HMI tags "xDI"
   "DIx_DB_M1_QF_Input" : Bool = PLC DIx_DB.M1_QF.Input AT %DB200.DBX0.0, 1 s
   "DIx_DB_M1_QF_Signal" : Bool = PLC DIx_DB.M1_QF.Signal AT %DB200.DBX2.0, 1 s
   "DIx_DB_M1_QF_Hand" : Bool = PLC DIx_DB.M1_QF.Hand AT %DB200.DBX4.0, 1 s
   "DIx_DB_M1_QF_Start_M" : Bool = PLC DIx_DB.M1_QF.Start_M AT %DB200.DBX4.1, 1 s
   "DIx_DB_M1_QF_Inverse" : Bool = PLC DIx_DB.M1_QF.Inverse AT %DB200.DBX4.3, 1 s
   "DIx_DB_M1_QF_Filter_On_SP" : Int = PLC DIx_DB.M1_QF.Filter_On.SP AT %DB200.DBW6, 1 s
   "DIx_DB_M1_QF_Filter_Off_SP" : Int = PLC DIx_DB.M1_QF.Filter_Off.SP AT %DB200.DBW12, 1 s
   "DIx_DB_M2_QF_Input" : Bool = PLC DIx_DB.M2_QF.Input AT %DB200.DBX20.0, 1 s
   "DIx_DB_M2_QF_Signal" : Bool = PLC DIx_DB.M2_QF.Signal AT %DB200.DBX22.0, 1 s
   "DIx_DB_M2_QF_Hand" : Bool = PLC DIx_DB.M2_QF.Hand AT %DB200.DBX24.0, 1 s
   "DIx_DB_M2_QF_Start_M" : Bool = PLC DIx_DB.M2_QF.Start_M AT %DB200.DBX24.1, 1 s
   "DIx_DB_M2_QF_Inverse" : Bool = PLC DIx_DB.M2_QF.Inverse AT %DB200.DBX24.3, 1 s
   "DIx_DB_M2_QF_Filter_On_SP" : Int = PLC DIx_DB.M2_QF.Filter_On.SP AT %DB200.DBW26, 1 s
   "DIx_DB_M2_QF_Filter_Off_SP" : Int = PLC DIx_DB.M2_QF.Filter_Off.SP AT %DB200.DBW32, 1 s
   "DIx_DB_M3_QF_Input" : Bool = PLC DIx_DB.M3_QF.Input AT %DB200.DBX40.0, 1 s
   "DIx_DB_M3_QF_Signal" : Bool = PLC DIx_DB.M3_QF.Signal AT %DB200.DBX42.0, 1 s
   "DIx_DB_M3_QF_Hand" : Bool = PLC DIx_DB.M3_QF.Hand AT %DB200.DBX44.0, 1 s
   "DIx_DB_M3_QF_Start_M" : Bool = PLC DIx_DB.M3_QF.Start_M AT %DB200.DBX44.1, 1 s
   "DIx_DB_M3_QF_Inverse" : Bool = PLC DIx_DB.M3_QF.Inverse AT %DB200.DBX44.3, 1 s
   "DIx_DB_M3_QF_Filter_On_SP" : Int = PLC DIx_DB.M3_QF.Filter_On.SP AT %DB200.DBW46, 1 s
   "DIx_DB_M3_QF_Filter_Off_SP" : Int = PLC DIx_DB.M3_QF.Filter_Off.SP AT %DB200.DBW52, 1 s
   "DIx_DB_Heat_1_Input" : Bool = PLC DIx_DB.Heat_1.Input AT %DB200.DBX60.0, 1 s
   "DIx_DB_Heat_1_Signal" : Bool = PLC DIx_DB.Heat_1.Signal AT %DB200.DBX62.0, 1 s
   "DIx_DB_Heat_1_Hand" : Bool = PLC DIx_DB.Heat_1.Hand AT %DB200.DBX64.0, 1 s
   "DIx_DB_Heat_1_Start_M" : Bool = PLC DIx_DB.Heat_1.Start_M AT %DB200.DBX64.1, 1 s
   "DIx_DB_Heat_1_Filter_On_SP" : Int = PLC DIx_DB.Heat_1.Filter_On.SP AT %DB200.DBW66, 1 s
   "DIx_DB_Heat_1_Filter_Off_SP" : Int = PLC DIx_DB.Heat_1.Filter_Off.SP AT %DB200.DBW72, 1 s
   "DIx_DB_Heat_2_Filter_Off_SP" : Int = PLC DIx_DB.Heat_2.Filter_Off.SP AT %DB200.DBW92, 1 s
   "DIx_DB_Heat_2_Filter_On_SP" : Int = PLC DIx_DB.Heat_2.Filter_On.SP AT %DB200.DBW86, 1 s
   "DIx_DB_Heat_2_Inverse" : Bool = PLC DIx_DB.Heat_2.Inverse AT %DB200.DBX84.3, 1 s
   "DIx_DB_Heat_2_Start_M" : Bool = PLC DIx_DB.Heat_2.Start_M AT %DB200.DBX84.1, 1 s
   "DIx_DB_Heat_2_Hand" : Bool = PLC DIx_DB.Heat_2.Hand AT %DB200.DBX84.0, 1 s
   "DIx_DB_Heat_2_Signal" : Bool = PLC DIx_DB.Heat_2.Signal AT %DB200.DBX82.0, 1 s
   "DIx_DB_Heat_2_Input" : Bool = PLC DIx_DB.Heat_2.Input AT %DB200.DBX80.0, 1 s
   "DIx_DB_Heat_3_Input" : Bool = PLC DIx_DB.Heat_3.Input AT %DB200.DBX100.0, 1 s
   "DIx_DB_Heat_3_Signal" : Bool = PLC DIx_DB.Heat_3.Signal AT %DB200.DBX102.0, 1 s
   "DIx_DB_Heat_3_Hand" : Bool = PLC DIx_DB.Heat_3.Hand AT %DB200.DBX104.0, 1 s
   "DIx_DB_Heat_3_Start_M" : Bool = PLC DIx_DB.Heat_3.Start_M AT %DB200.DBX104.1, 1 s
   "DIx_DB_Heat_3_Inverse" : Bool = PLC DIx_DB.Heat_3.Inverse AT %DB200.DBX104.3, 1 s
   "DIx_DB_Heat_3_Filter_Off_SP" : Int = PLC DIx_DB.Heat_3.Filter_Off.SP AT %DB200.DBW112, 1 s
   "DIx_DB_Heat_3_Filter_On_SP" : Int = PLC DIx_DB.Heat_3.Filter_On.SP AT %DB200.DBW106, 1 s
   "DIx_DB_AllBlock_Input" : Bool = PLC DIx_DB.AllBlock.Input AT %DB200.DBX140.0, 1 s
   "DIx_DB_AllBlock_Signal" : Bool = PLC DIx_DB.AllBlock.Signal AT %DB200.DBX142.0, 1 s
   "DIx_DB_AllBlock_Hand" : Bool = PLC DIx_DB.AllBlock.Hand AT %DB200.DBX144.0, 1 s
   "DIx_DB_AllBlock_Start_M" : Bool = PLC DIx_DB.AllBlock.Start_M AT %DB200.DBX144.1, 1 s
   "DIx_DB_AllBlock_Inverse" : Bool = PLC DIx_DB.AllBlock.Inverse AT %DB200.DBX144.3, 1 s
   "DIx_DB_AllBlock_Filter_On_SP" : Int = PLC DIx_DB.AllBlock.Filter_On.SP AT %DB200.DBW146, 1 s
   "DIx_DB_AllBlock_Filter_Off_SP" : Int = PLC DIx_DB.AllBlock.Filter_Off.SP AT %DB200.DBW152, 1 s
   "DIx_DB_Mass_1_Input" : Bool = PLC DIx_DB.Mass_1.Input AT %DB200.DBX160.0, 1 s
   "DIx_DB_Mass_1_Signal" : Bool = PLC DIx_DB.Mass_1.Signal AT %DB200.DBX162.0, 1 s
   "DIx_DB_Mass_1_Hand" : Bool = PLC DIx_DB.Mass_1.Hand AT %DB200.DBX164.0, 1 s
   "DIx_DB_Mass_1_Start_M" : Bool = PLC DIx_DB.Mass_1.Start_M AT %DB200.DBX164.1, 1 s
   "DIx_DB_Mass_1_Inverse" : Bool = PLC DIx_DB.Mass_1.Inverse AT %DB200.DBX164.3, 1 s
   "DIx_DB_Mass_1_Filter_On_SP" : Int = PLC DIx_DB.Mass_1.Filter_On.SP AT %DB200.DBW166, 1 s
   "DIx_DB_Mass_1_Filter_Off_SP" : Int = PLC DIx_DB.Mass_1.Filter_Off.SP AT %DB200.DBW172, 1 s
   "DIx_DB_Mass_2_Input" : Bool = PLC DIx_DB.Mass_2.Input AT %DB200.DBX180.0, 1 s
   "DIx_DB_Mass_2_Signal" : Bool = PLC DIx_DB.Mass_2.Signal AT %DB200.DBX182.0, 1 s
   "DIx_DB_Mass_2_Hand" : Bool = PLC DIx_DB.Mass_2.Hand AT %DB200.DBX184.0, 1 s
   "DIx_DB_Mass_2_Start_M" : Bool = PLC DIx_DB.Mass_2.Start_M AT %DB200.DBX184.1, 1 s
   "DIx_DB_Mass_2_Inverse" : Bool = PLC DIx_DB.Mass_2.Inverse AT %DB200.DBX184.3, 1 s
   "DIx_DB_Mass_2_Filter_On_SP" : Int = PLC DIx_DB.Mass_2.Filter_On.SP AT %DB200.DBW186, 1 s
   "DIx_DB_Mass_2_Filter_Off_SP" : Int = PLC DIx_DB.Mass_2.Filter_Off.SP AT %DB200.DBW192, 1 s
   "DIx_DB_Heat_4_Hand" : Bool = PLC DIx_DB.Heat_4.Hand AT %DB200.DBX124.0, 1 s
   "DIx_DB_Heat_4_Start_M" : Bool = PLC DIx_DB.Heat_4.Start_M AT %DB200.DBX124.1, 1 s
   "DIx_DB_Heat_4_Inverse" : Bool = PLC DIx_DB.Heat_4.Inverse AT %DB200.DBX124.3, 1 s
   "DIx_DB_Heat_4_Filter_On_SP" : Int = PLC DIx_DB.Heat_4.Filter_On.SP AT %DB200.DBW126, 1 s
   "DIx_DB_Heat_4_Filter_Off_SP" : Int = PLC DIx_DB.Heat_4.Filter_Off.SP AT %DB200.DBW132, 1 s

HMI tags "xDO"
   "DOx_DB_M1_CMD_Start_A" : Bool = PLC DOx_DB.M1_CMD.Start_A AT %DB201.DBX0.0, 1 s
   "DOx_DB_M1_CMD_Q" : Bool = PLC DOx_DB.M1_CMD.Q AT %DB201.DBX0.2, 1 s
   "DOx_DB_M1_CMD_Hand" : Bool = PLC DOx_DB.M1_CMD.Hand AT %DB201.DBX2.0, 1 s
   "DOx_DB_M1_CMD_Start_M" : Bool = PLC DOx_DB.M1_CMD.Start_M AT %DB201.DBX2.1, 1 s
   "DOx_DB_M1_CMD_Simulation" : Bool = PLC DOx_DB.M1_CMD.Simulation AT %DB201.DBX2.2, 1 s
   "DOx_DB_M1_CMD_Inverse" : Bool = PLC DOx_DB.M1_CMD.Inverse AT %DB201.DBX2.3, 1 s
   "DOx_DB_M2_CMD_Start_A" : Bool = PLC DOx_DB.M2_CMD.Start_A AT %DB201.DBX10.0, 1 s
   "DOx_DB_M2_CMD_Q" : Bool = PLC DOx_DB.M2_CMD.Q AT %DB201.DBX10.2, 1 s
   "DOx_DB_M2_CMD_Hand" : Bool = PLC DOx_DB.M2_CMD.Hand AT %DB201.DBX12.0, 1 s
   "DOx_DB_M2_CMD_Start_M" : Bool = PLC DOx_DB.M2_CMD.Start_M AT %DB201.DBX12.1, 1 s
   "DOx_DB_M2_CMD_Simulation" : Bool = PLC DOx_DB.M2_CMD.Simulation AT %DB201.DBX12.2, 1 s
   "DOx_DB_M2_CMD_Inverse" : Bool = PLC DOx_DB.M2_CMD.Inverse AT %DB201.DBX12.3, 1 s
   "DOx_DB_M3_CMD_Start_A" : Bool = PLC DOx_DB.M3_CMD.Start_A AT %DB201.DBX20.0, 1 s
   "DOx_DB_M3_CMD_Q" : Bool = PLC DOx_DB.M3_CMD.Q AT %DB201.DBX20.2, 1 s
   "DOx_DB_M3_CMD_Hand" : Bool = PLC DOx_DB.M3_CMD.Hand AT %DB201.DBX22.0, 1 s
   "DOx_DB_M3_CMD_Start_M" : Bool = PLC DOx_DB.M3_CMD.Start_M AT %DB201.DBX22.1, 1 s
   "DOx_DB_M3_CMD_Simulation" : Bool = PLC DOx_DB.M3_CMD.Simulation AT %DB201.DBX22.2, 1 s
   "DOx_DB_M3_CMD_Inverse" : Bool = PLC DOx_DB.M3_CMD.Inverse AT %DB201.DBX22.3, 1 s
   "DOx_DB_LED_Error_1_Start_A" : Bool = PLC DOx_DB.LED_Error_1.Start_A AT %DB201.DBX30.0, 1 s
   "DOx_DB_LED_Error_1_Q" : Bool = PLC DOx_DB.LED_Error_1.Q AT %DB201.DBX30.2, 1 s
   "DOx_DB_LED_Error_1_Hand" : Bool = PLC DOx_DB.LED_Error_1.Hand AT %DB201.DBX32.0, 1 s
   "DOx_DB_LED_Error_1_Simulation" : Bool = PLC DOx_DB.LED_Error_1.Simulation AT %DB201.DBX32.2, 1 s
   "DOx_DB_LED_Error_1_Start_M" : Bool = PLC DOx_DB.LED_Error_1.Start_M AT %DB201.DBX32.1, 1 s
   "DOx_DB_LED_Error_1_Inverse" : Bool = PLC DOx_DB.LED_Error_1.Inverse AT %DB201.DBX32.3, 1 s
   "DOx_DB_LED_Error_2_Start_A" : Bool = PLC DOx_DB.LED_Error_2.Start_A AT %DB201.DBX40.0, 1 s
   "DOx_DB_LED_Error_2_Q" : Bool = PLC DOx_DB.LED_Error_2.Q AT %DB201.DBX40.2, 1 s
   "DOx_DB_LED_Error_2_Hand" : Bool = PLC DOx_DB.LED_Error_2.Hand AT %DB201.DBX42.0, 1 s
   "DOx_DB_LED_Error_2_Start_M" : Bool = PLC DOx_DB.LED_Error_2.Start_M AT %DB201.DBX42.1, 1 s
   "DOx_DB_LED_Error_2_Simulation" : Bool = PLC DOx_DB.LED_Error_2.Simulation AT %DB201.DBX42.2, 1 s
   "DOx_DB_LED_Error_2_Inverse" : Bool = PLC DOx_DB.LED_Error_2.Inverse AT %DB201.DBX42.3, 1 s
   "DOx_DB_LED_Alarm_Start_A" : Bool = PLC DOx_DB.LED_Alarm.Start_A AT %DB201.DBX50.0, 1 s
   "DOx_DB_LED_Alarm_Q" : Bool = PLC DOx_DB.LED_Alarm.Q AT %DB201.DBX50.2, 1 s
   "DOx_DB_LED_Alarm_Hand" : Bool = PLC DOx_DB.LED_Alarm.Hand AT %DB201.DBX52.0, 1 s
   "DOx_DB_LED_Alarm_Start_M" : Bool = PLC DOx_DB.LED_Alarm.Start_M AT %DB201.DBX52.1, 1 s
   "DOx_DB_LED_Alarm_Simulation" : Bool = PLC DOx_DB.LED_Alarm.Simulation AT %DB201.DBX52.2, 1 s
   "DOx_DB_LED_Alarm_Inverse" : Bool = PLC DOx_DB.LED_Alarm.Inverse AT %DB201.DBX52.3, 1 s
   "DOx_DB_LED_M1_Alarm_Start_A" : Bool = PLC DOx_DB.LED_M1_Alarm.Start_A AT %DB201.DBX60.0, 1 s
   "DOx_DB_LED_M1_Alarm_Q" : Bool = PLC DOx_DB.LED_M1_Alarm.Q AT %DB201.DBX60.2, 1 s
   "DOx_DB_LED_M1_Alarm_Hand" : Bool = PLC DOx_DB.LED_M1_Alarm.Hand AT %DB201.DBX62.0, 1 s
   "DOx_DB_LED_M1_Alarm_Start_M" : Bool = PLC DOx_DB.LED_M1_Alarm.Start_M AT %DB201.DBX62.1, 1 s
   "DOx_DB_LED_M1_Alarm_Simulation" : Bool = PLC DOx_DB.LED_M1_Alarm.Simulation AT %DB201.DBX62.2, 1 s
   "DOx_DB_LED_M1_Alarm_Inverse" : Bool = PLC DOx_DB.LED_M1_Alarm.Inverse AT %DB201.DBX62.3, 1 s
   "DOx_DB_LED_M2_Alarm_Start_A" : Bool = PLC DOx_DB.LED_M2_Alarm.Start_A AT %DB201.DBX70.0, 1 s
   "DOx_DB_LED_M2_Alarm_Q" : Bool = PLC DOx_DB.LED_M2_Alarm.Q AT %DB201.DBX70.2, 1 s
   "DOx_DB_LED_M2_Alarm_Hand" : Bool = PLC DOx_DB.LED_M2_Alarm.Hand AT %DB201.DBX72.0, 1 s
   "DOx_DB_LED_M2_Alarm_Start_M" : Bool = PLC DOx_DB.LED_M2_Alarm.Start_M AT %DB201.DBX72.1, 1 s
   "DOx_DB_LED_M2_Alarm_Simulation" : Bool = PLC DOx_DB.LED_M2_Alarm.Simulation AT %DB201.DBX72.2, 1 s
   "DOx_DB_LED_M2_Alarm_Inverse" : Bool = PLC DOx_DB.LED_M2_Alarm.Inverse AT %DB201.DBX72.3, 1 s
   "DOx_DB_LED_M3_Alarm_Start_A" : Bool = PLC DOx_DB.LED_M3_Alarm.Start_A AT %DB201.DBX80.0, 1 s
   "DOx_DB_LED_M3_Alarm_Q" : Bool = PLC DOx_DB.LED_M3_Alarm.Q AT %DB201.DBX80.2, 1 s
   "DOx_DB_LED_M3_Alarm_Hand" : Bool = PLC DOx_DB.LED_M3_Alarm.Hand AT %DB201.DBX82.0, 1 s
   "DOx_DB_LED_M3_Alarm_Start_M" : Bool = PLC DOx_DB.LED_M3_Alarm.Start_M AT %DB201.DBX82.1, 1 s
   "DOx_DB_LED_M3_Alarm_Simulation" : Bool = PLC DOx_DB.LED_M3_Alarm.Simulation AT %DB201.DBX82.2, 1 s
   "DOx_DB_LED_M3_Alarm_Inverse" : Bool = PLC DOx_DB.LED_M3_Alarm.Inverse AT %DB201.DBX82.3, 1 s

HMI tags "xAI"
   "AIx_DB_Flow_1_Signal" : Int = PLC AIx_DB.Flow_1.Signal AT %DB202.DBW0, 1 s
   "AIx_DB_Flow_1_Result" : Real = PLC AIx_DB.Flow_1.Result AT %DB202.DBD6, 1 s
   "AIx_DB_Flow_1_CMD_Start_A" : Bool = PLC AIx_DB.Flow_1.CMD.Start_A AT %DB202.DBX10.1, 1 s
   "AIx_DB_Flow_1_CMD_Hand" : Bool = PLC AIx_DB.Flow_1.CMD.Hand AT %DB202.DBX10.0, 1 s
   "AIx_DB_Flow_1_Use_RTD" : Bool = PLC AIx_DB.Flow_1.Use.RTD AT %DB202.DBX16.0, 1 s
   "AIx_DB_Flow_1_Use_Filter" : Bool = PLC AIx_DB.Flow_1.Use.Filter AT %DB202.DBX16.1, 1 s
   "AIx_DB_Flow_1_RTD_c" : Real = PLC AIx_DB.Flow_1.RTD_c AT %DB202.DBD30, 1 s
   "AIx_DB_Flow_1_Calibration" : Real = PLC AIx_DB.Flow_1.Calibration AT %DB202.DBD34, 1 s
   "AIx_DB_Flow_1_Converter_Min_In" : Real = PLC AIx_DB.Flow_1.Converter.Min_In AT %DB202.DBD60, 1 s
   "AIx_DB_Flow_1_Converter_Max_In" : Real = PLC AIx_DB.Flow_1.Converter.Max_In AT %DB202.DBD64, 1 s
   "AIx_DB_Flow_1_Converter_Min_Out" : Real = PLC AIx_DB.Flow_1.Converter.Min_Out AT %DB202.DBD68, 1 s
   "AIx_DB_Flow_1_Converter_Max_Out" : Real = PLC AIx_DB.Flow_1.Converter.Max_Out AT %DB202.DBD72, 1 s
   "AIx_DB_Flow_1_Filter_SP" : Real = PLC AIx_DB.Flow_1.Filter.SP AT %DB202.DBD38, 1 s
   "AIx_DB_Flow_1_SP_NC" : Real = PLC AIx_DB.Flow_1.SP.NC AT %DB202.DBD76, 1 s
   "AIx_DB_Flow_1_SP_SC" : Real = PLC AIx_DB.Flow_1.SP.SC AT %DB202.DBD80, 1 s
   "AIx_DB_Flow_1_SP_HH" : Real = PLC AIx_DB.Flow_1.SP.HH AT %DB202.DBD84, 1 s
   "AIx_DB_Flow_1_SP_H" : Real = PLC AIx_DB.Flow_1.SP.H AT %DB202.DBD88, 1 s
   "AIx_DB_Flow_1_SP_L" : Real = PLC AIx_DB.Flow_1.SP.L AT %DB202.DBD92, 1 s
   "AIx_DB_Flow_1_SP_LL" : Real = PLC AIx_DB.Flow_1.SP.LL AT %DB202.DBD96, 1 s
   "AIx_DB_Flow_1_Alarm" : Word = PLC AIx_DB.Flow_1.Alarm AT %DB202.DBW138, 1 s
   "AIx_DB_Flow_1_Timers_NC_SP" : Int = PLC AIx_DB.Flow_1.Timers.NC.SP AT %DB202.DBW100, 1 s
   "AIx_DB_Flow_1_Timers_SC_SP" : Int = PLC AIx_DB.Flow_1.Timers.SC.SP AT %DB202.DBW106, 1 s
   "AIx_DB_Flow_1_Timers_HH_SP" : Int = PLC AIx_DB.Flow_1.Timers.HH.SP AT %DB202.DBW112, 1 s
   "AIx_DB_Flow_1_Timers_H_SP" : Int = PLC AIx_DB.Flow_1.Timers.H.SP AT %DB202.DBW118, 1 s
   "AIx_DB_Flow_1_Timers_L_SP" : Int = PLC AIx_DB.Flow_1.Timers.L.SP AT %DB202.DBW124, 1 s
   "AIx_DB_Flow_1_Timers_LL_SP" : Int = PLC AIx_DB.Flow_1.Timers.LL.SP AT %DB202.DBW130, 1 s
   "AIx_DB_Flow_2_Signal" : Int = PLC AIx_DB.Flow_2.Signal AT %DB202.DBW140, 1 s
   "AIx_DB_Flow_2_Result" : Real = PLC AIx_DB.Flow_2.Result AT %DB202.DBD146, 1 s
   "AIx_DB_Flow_2_CMD_Start_A" : Bool = PLC AIx_DB.Flow_2.CMD.Start_A AT %DB202.DBX150.1, 1 s
   "AIx_DB_Flow_2_CMD_Hand" : Bool = PLC AIx_DB.Flow_2.CMD.Hand AT %DB202.DBX150.0, 1 s
   "AIx_DB_Flow_2_Use_RTD" : Bool = PLC AIx_DB.Flow_2.Use.RTD AT %DB202.DBX156.0, 1 s
   "AIx_DB_Flow_2_Use_Filter" : Bool = PLC AIx_DB.Flow_2.Use.Filter AT %DB202.DBX156.1, 1 s
   "AIx_DB_Flow_2_RTD_c" : Real = PLC AIx_DB.Flow_2.RTD_c AT %DB202.DBD170, 1 s
   "AIx_DB_Flow_2_Calibration" : Real = PLC AIx_DB.Flow_2.Calibration AT %DB202.DBD174, 1 s
   "AIx_DB_Flow_2_Converter_Min_In" : Real = PLC AIx_DB.Flow_2.Converter.Min_In AT %DB202.DBD200, 1 s
   "AIx_DB_Flow_2_Converter_Max_In" : Real = PLC AIx_DB.Flow_2.Converter.Max_In AT %DB202.DBD204, 1 s
   "AIx_DB_Flow_2_Converter_Min_Out" : Real = PLC AIx_DB.Flow_2.Converter.Min_Out AT %DB202.DBD208, 1 s
   "AIx_DB_Flow_2_Converter_Max_Out" : Real = PLC AIx_DB.Flow_2.Converter.Max_Out AT %DB202.DBD212, 1 s
   "AIx_DB_Flow_2_Filter_SP" : Real = PLC AIx_DB.Flow_2.Filter.SP AT %DB202.DBD178, 1 s
   "AIx_DB_Flow_2_SP_NC" : Real = PLC AIx_DB.Flow_2.SP.NC AT %DB202.DBD216, 1 s
   "AIx_DB_Flow_2_SP_SC" : Real = PLC AIx_DB.Flow_2.SP.SC AT %DB202.DBD220, 1 s
   "AIx_DB_Flow_2_SP_HH" : Real = PLC AIx_DB.Flow_2.SP.HH AT %DB202.DBD224, 1 s
   "AIx_DB_Flow_2_SP_H" : Real = PLC AIx_DB.Flow_2.SP.H AT %DB202.DBD228, 1 s
   "AIx_DB_Flow_2_SP_L" : Real = PLC AIx_DB.Flow_2.SP.L AT %DB202.DBD232, 1 s
   "AIx_DB_Flow_2_SP_LL" : Real = PLC AIx_DB.Flow_2.SP.LL AT %DB202.DBD236, 1 s
   "AIx_DB_Flow_2_Alarm" : Word = PLC AIx_DB.Flow_2.Alarm AT %DB202.DBW278, 1 s
   "AIx_DB_Flow_2_Timers_NC_SP" : Int = PLC AIx_DB.Flow_2.Timers.NC.SP AT %DB202.DBW240, 1 s
   "AIx_DB_Flow_2_Timers_SC_SP" : Int = PLC AIx_DB.Flow_2.Timers.SC.SP AT %DB202.DBW246, 1 s
   "AIx_DB_Flow_2_Timers_HH_SP" : Int = PLC AIx_DB.Flow_2.Timers.HH.SP AT %DB202.DBW252, 1 s
   "AIx_DB_Flow_2_Timers_H_SP" : Int = PLC AIx_DB.Flow_2.Timers.H.SP AT %DB202.DBW258, 1 s
   "AIx_DB_Flow_2_Timers_L_SP" : Int = PLC AIx_DB.Flow_2.Timers.L.SP AT %DB202.DBW264, 1 s
   "AIx_DB_Flow_2_Timers_LL_SP" : Int = PLC AIx_DB.Flow_2.Timers.LL.SP AT %DB202.DBW270, 1 s
   "AIx_DB_Trans_1_Signal" : Int = PLC AIx_DB.Trans_1.Signal AT %DB202.DBW280, 1 s
   "AIx_DB_Trans_1_Result" : Real = PLC AIx_DB.Trans_1.Result AT %DB202.DBD286, 1 s
   "AIx_DB_Trans_1_CMD_Start_A" : Bool = PLC AIx_DB.Trans_1.CMD.Start_A AT %DB202.DBX290.1, 1 s
   "AIx_DB_Trans_1_CMD_Hand" : Bool = PLC AIx_DB.Trans_1.CMD.Hand AT %DB202.DBX290.0, 1 s
   "AIx_DB_Trans_1_Use_RTD" : Bool = PLC AIx_DB.Trans_1.Use.RTD AT %DB202.DBX296.0, 1 s
   "AIx_DB_Trans_1_Use_Filter" : Bool = PLC AIx_DB.Trans_1.Use.Filter AT %DB202.DBX296.1, 1 s
   "AIx_DB_Trans_1_RTD_c" : Real = PLC AIx_DB.Trans_1.RTD_c AT %DB202.DBD310, 1 s
   "AIx_DB_Trans_1_Calibration" : Real = PLC AIx_DB.Trans_1.Calibration AT %DB202.DBD314, 1 s
   "AIx_DB_Trans_1_Converter_Min_In" : Real = PLC AIx_DB.Trans_1.Converter.Min_In AT %DB202.DBD340, 1 s
   "AIx_DB_Trans_1_Converter_Max_In" : Real = PLC AIx_DB.Trans_1.Converter.Max_In AT %DB202.DBD344, 1 s
   "AIx_DB_Trans_1_Converter_Min_Out" : Real = PLC AIx_DB.Trans_1.Converter.Min_Out AT %DB202.DBD348, 1 s
   "AIx_DB_Trans_1_Converter_Max_Out" : Real = PLC AIx_DB.Trans_1.Converter.Max_Out AT %DB202.DBD352, 1 s
   "AIx_DB_Trans_1_Filter_SP" : Real = PLC AIx_DB.Trans_1.Filter.SP AT %DB202.DBD318, 1 s
   "AIx_DB_Trans_1_SP_NC" : Real = PLC AIx_DB.Trans_1.SP.NC AT %DB202.DBD356, 1 s
   "AIx_DB_Trans_1_SP_SC" : Real = PLC AIx_DB.Trans_1.SP.SC AT %DB202.DBD360, 1 s
   "AIx_DB_Trans_1_SP_HH" : Real = PLC AIx_DB.Trans_1.SP.HH AT %DB202.DBD364, 1 s
   "AIx_DB_Trans_1_SP_H" : Real = PLC AIx_DB.Trans_1.SP.H AT %DB202.DBD368, 1 s
   "AIx_DB_Trans_1_SP_L" : Real = PLC AIx_DB.Trans_1.SP.L AT %DB202.DBD372, 1 s
   "AIx_DB_Trans_1_SP_LL" : Real = PLC AIx_DB.Trans_1.SP.LL AT %DB202.DBD376, 1 s
   "AIx_DB_Trans_1_Alarm" : Word = PLC AIx_DB.Trans_1.Alarm AT %DB202.DBW418, 1 s
   "AIx_DB_Trans_1_Timers_NC_SP" : Int = PLC AIx_DB.Trans_1.Timers.NC.SP AT %DB202.DBW380, 1 s
   "AIx_DB_Trans_1_Timers_SC_SP" : Int = PLC AIx_DB.Trans_1.Timers.SC.SP AT %DB202.DBW386, 1 s
   "AIx_DB_Trans_1_Timers_HH_SP" : Int = PLC AIx_DB.Trans_1.Timers.HH.SP AT %DB202.DBW392, 1 s
   "AIx_DB_Trans_1_Timers_H_SP" : Int = PLC AIx_DB.Trans_1.Timers.H.SP AT %DB202.DBW398, 1 s
   "AIx_DB_Trans_1_Timers_L_SP" : Int = PLC AIx_DB.Trans_1.Timers.L.SP AT %DB202.DBW404, 1 s
   "AIx_DB_Trans_1_Timers_LL_SP" : Int = PLC AIx_DB.Trans_1.Timers.LL.SP AT %DB202.DBW410, 1 s
   "AIx_DB_Trans_2_Signal" : Int = PLC AIx_DB.Trans_2.Signal AT %DB202.DBW420, 1 s
   "AIx_DB_Trans_2_Result" : Real = PLC AIx_DB.Trans_2.Result AT %DB202.DBD426, 1 s
   "AIx_DB_Trans_2_CMD_Start_A" : Bool = PLC AIx_DB.Trans_2.CMD.Start_A AT %DB202.DBX430.1, 1 s
   "AIx_DB_Trans_2_CMD_Hand" : Bool = PLC AIx_DB.Trans_2.CMD.Hand AT %DB202.DBX430.0, 1 s
   "AIx_DB_Trans_2_Use_RTD" : Bool = PLC AIx_DB.Trans_2.Use.RTD AT %DB202.DBX436.0, 1 s
   "AIx_DB_Trans_2_Use_Filter" : Bool = PLC AIx_DB.Trans_2.Use.Filter AT %DB202.DBX436.1, 1 s
   "AIx_DB_Trans_2_RTD_c" : Real = PLC AIx_DB.Trans_2.RTD_c AT %DB202.DBD450, 1 s
   "AIx_DB_Trans_2_Calibration" : Real = PLC AIx_DB.Trans_2.Calibration AT %DB202.DBD454, 1 s
   "AIx_DB_Trans_2_Converter_Min_In" : Real = PLC AIx_DB.Trans_2.Converter.Min_In AT %DB202.DBD480, 1 s
   "AIx_DB_Trans_2_Converter_Max_In" : Real = PLC AIx_DB.Trans_2.Converter.Max_In AT %DB202.DBD484, 1 s
   "AIx_DB_Trans_2_Converter_Min_Out" : Real = PLC AIx_DB.Trans_2.Converter.Min_Out AT %DB202.DBD488, 1 s
   "AIx_DB_Trans_2_Converter_Max_Out" : Real = PLC AIx_DB.Trans_2.Converter.Max_Out AT %DB202.DBD492, 1 s
   "AIx_DB_Trans_2_Filter_SP" : Real = PLC AIx_DB.Trans_2.Filter.SP AT %DB202.DBD458, 1 s
   "AIx_DB_Trans_2_SP_NC" : Real = PLC AIx_DB.Trans_2.SP.NC AT %DB202.DBD496, 1 s
   "AIx_DB_Trans_2_SP_SC" : Real = PLC AIx_DB.Trans_2.SP.SC AT %DB202.DBD500, 1 s
   "AIx_DB_Trans_2_SP_HH" : Real = PLC AIx_DB.Trans_2.SP.HH AT %DB202.DBD504, 1 s
   "AIx_DB_Trans_2_SP_H" : Real = PLC AIx_DB.Trans_2.SP.H AT %DB202.DBD508, 1 s
   "AIx_DB_Trans_2_SP_L" : Real = PLC AIx_DB.Trans_2.SP.L AT %DB202.DBD512, 1 s
   "AIx_DB_Trans_2_SP_LL" : Real = PLC AIx_DB.Trans_2.SP.LL AT %DB202.DBD516, 1 s
   "AIx_DB_Trans_2_Alarm" : Word = PLC AIx_DB.Trans_2.Alarm AT %DB202.DBW558, 1 s
   "AIx_DB_Trans_2_Timers_NC_SP" : Int = PLC AIx_DB.Trans_2.Timers.NC.SP AT %DB202.DBW520, 1 s
   "AIx_DB_Trans_2_Timers_SC_SP" : Int = PLC AIx_DB.Trans_2.Timers.SC.SP AT %DB202.DBW526, 1 s
   "AIx_DB_Trans_2_Timers_HH_SP" : Int = PLC AIx_DB.Trans_2.Timers.HH.SP AT %DB202.DBW532, 1 s
   "AIx_DB_Trans_2_Timers_H_SP" : Int = PLC AIx_DB.Trans_2.Timers.H.SP AT %DB202.DBW538, 1 s
   "AIx_DB_Trans_2_Timers_L_SP" : Int = PLC AIx_DB.Trans_2.Timers.L.SP AT %DB202.DBW544, 1 s
   "AIx_DB_Trans_2_Timers_LL_SP" : Int = PLC AIx_DB.Trans_2.Timers.LL.SP AT %DB202.DBW550, 1 s
   "AIx_DB_Flow_3_Result" : Real = PLC AIx_DB.Flow_3.Result AT %DB202.DBD566, 1 s
   "AIx_DB_Flow_3_Signal" : Int = PLC AIx_DB.Flow_3.Signal AT %DB202.DBW560, 1 s
   "AIx_DB_Flow_3_CMD_Hand" : Bool = PLC AIx_DB.Flow_3.CMD.Hand AT %DB202.DBX570.0, 1 s
   "AIx_DB_Flow_3_CMD_Start_A" : Bool = PLC AIx_DB.Flow_3.CMD.Start_A AT %DB202.DBX570.1, 1 s
   "AIx_DB_Flow_3_Use_RTD" : Bool = PLC AIx_DB.Flow_3.Use.RTD AT %DB202.DBX576.0, 1 s
   "AIx_DB_Flow_3_Use_Filter" : Bool = PLC AIx_DB.Flow_3.Use.Filter AT %DB202.DBX576.1, 1 s
   "AIx_DB_Flow_3_RTD_c" : Real = PLC AIx_DB.Flow_3.RTD_c AT %DB202.DBD590, 1 s
   "AIx_DB_Flow_3_SP_NC" : Real = PLC AIx_DB.Flow_3.SP.NC AT %DB202.DBD636, 1 s
   "AIx_DB_Flow_3_SP_LL" : Real = PLC AIx_DB.Flow_3.SP.LL AT %DB202.DBD656, 1 s
   "AIx_DB_Flow_3_SP_L" : Real = PLC AIx_DB.Flow_3.SP.L AT %DB202.DBD652, 1 s
   "AIx_DB_Flow_3_SP_H" : Real = PLC AIx_DB.Flow_3.SP.H AT %DB202.DBD648, 1 s
   "AIx_DB_Flow_3_SP_HH" : Real = PLC AIx_DB.Flow_3.SP.HH AT %DB202.DBD644, 1 s
   "AIx_DB_Flow_3_SP_SC" : Real = PLC AIx_DB.Flow_3.SP.SC AT %DB202.DBD640, 1 s
   "AIx_DB_Flow_3_Timers_NC_SP" : Int = PLC AIx_DB.Flow_3.Timers.NC.SP AT %DB202.DBW660, 1 s
   "AIx_DB_Flow_3_Timers_SC_SP" : Int = PLC AIx_DB.Flow_3.Timers.SC.SP AT %DB202.DBW666, 1 s
   "AIx_DB_Flow_3_Timers_HH_SP" : Int = PLC AIx_DB.Flow_3.Timers.HH.SP AT %DB202.DBW672, 1 s
   "AIx_DB_Flow_3_Timers_H_SP" : Int = PLC AIx_DB.Flow_3.Timers.H.SP AT %DB202.DBW678, 1 s
   "AIx_DB_Flow_3_Timers_L_SP" : Int = PLC AIx_DB.Flow_3.Timers.L.SP AT %DB202.DBW684, 1 s
   "AIx_DB_Flow_3_Timers_LL_SP" : Int = PLC AIx_DB.Flow_3.Timers.LL.SP AT %DB202.DBW690, 1 s
   "AIx_DB_Flow_3_Filter_SP" : Real = PLC AIx_DB.Flow_3.Filter.SP AT %DB202.DBD598, 1 s
   "AIx_DB_Flow_4_Timers_LL_SP" : Int = PLC AIx_DB.Flow_4.Timers.LL.SP AT %DB202.DBW830, 1 s
   "AIx_DB_Flow_4_Timers_L_SP" : Int = PLC AIx_DB.Flow_4.Timers.L.SP AT %DB202.DBW824, 1 s
   "AIx_DB_Flow_4_Timers_H_SP" : Int = PLC AIx_DB.Flow_4.Timers.H.SP AT %DB202.DBW818, 1 s
   "AIx_DB_Flow_4_Timers_HH_SP" : Int = PLC AIx_DB.Flow_4.Timers.HH.SP AT %DB202.DBW812, 1 s
   "AIx_DB_Flow_4_Timers_SC_SP" : Int = PLC AIx_DB.Flow_4.Timers.SC.SP AT %DB202.DBW806, 1 s
   "AIx_DB_Flow_4_Timers_NC_SP" : Int = PLC AIx_DB.Flow_4.Timers.NC.SP AT %DB202.DBW800, 1 s
   "AIx_DB_Flow_4_SP_NC" : Real = PLC AIx_DB.Flow_4.SP.NC AT %DB202.DBD776, 1 s
   "AIx_DB_Flow_4_SP_SC" : Real = PLC AIx_DB.Flow_4.SP.SC AT %DB202.DBD780, 1 s
   "AIx_DB_Flow_4_SP_HH" : Real = PLC AIx_DB.Flow_4.SP.HH AT %DB202.DBD784, 1 s
   "AIx_DB_Flow_4_SP_H" : Real = PLC AIx_DB.Flow_4.SP.H AT %DB202.DBD788, 1 s
   "AIx_DB_Flow_4_SP_L" : Real = PLC AIx_DB.Flow_4.SP.L AT %DB202.DBD792, 1 s
   "AIx_DB_Flow_4_SP_LL" : Real = PLC AIx_DB.Flow_4.SP.LL AT %DB202.DBD796, 1 s
   "AIx_DB_Flow_4_Converter_Max_Out" : Real = PLC AIx_DB.Flow_4.Converter.Max_Out AT %DB202.DBD772, 1 s
   "AIx_DB_Flow_4_Converter_Min_Out" : Real = PLC AIx_DB.Flow_4.Converter.Min_Out AT %DB202.DBD768, 1 s
   "AIx_DB_Flow_4_Converter_Max_In" : Real = PLC AIx_DB.Flow_4.Converter.Max_In AT %DB202.DBD764, 1 s
   "AIx_DB_Flow_4_Converter_Min_In" : Real = PLC AIx_DB.Flow_4.Converter.Min_In AT %DB202.DBD760, 1 s
   "AIx_DB_Flow_4_Filter_SP" : Real = PLC AIx_DB.Flow_4.Filter.SP AT %DB202.DBD738, 1 s
   "AIx_DB_Flow_4_RTD_c" : Real = PLC AIx_DB.Flow_4.RTD_c AT %DB202.DBD730, 1 s
   "AIx_DB_Flow_4_Use_RTD" : Bool = PLC AIx_DB.Flow_4.Use.RTD AT %DB202.DBX716.0, 1 s
   "AIx_DB_Flow_4_Use_Filter" : Bool = PLC AIx_DB.Flow_4.Use.Filter AT %DB202.DBX716.1, 1 s
   "AIx_DB_Flow_4_CMD_Hand" : Bool = PLC AIx_DB.Flow_4.CMD.Hand AT %DB202.DBX710.0, 1 s
   "AIx_DB_Flow_4_CMD_Start_A" : Bool = PLC AIx_DB.Flow_4.CMD.Start_A AT %DB202.DBX710.1, 1 s
   "AIx_DB_Flow_4_Result" : Real = PLC AIx_DB.Flow_4.Result AT %DB202.DBD706, 1 s
   "AIx_DB_Flow_4_Signal" : Int = PLC AIx_DB.Flow_4.Signal AT %DB202.DBW700, 1 s
   "AIx_DB_Flow_3_Converter_Max_Out" : Real = PLC AIx_DB.Flow_3.Converter.Max_Out AT %DB202.DBD632, 1 s
   "AIx_DB_Flow_3_Converter_Min_Out" : Real = PLC AIx_DB.Flow_3.Converter.Min_Out AT %DB202.DBD628, 1 s
   "AIx_DB_Flow_3_Converter_Max_In" : Real = PLC AIx_DB.Flow_3.Converter.Max_In AT %DB202.DBD624, 1 s
   "AIx_DB_Flow_3_Converter_Min_In" : Real = PLC AIx_DB.Flow_3.Converter.Min_In AT %DB202.DBD620, 1 s
   "AIx_DB_Flow_3_Calibration" : Real = PLC AIx_DB.Flow_3.Calibration AT %DB202.DBD594, 1 s
   "AIx_DB_Flow_4_Calibration" : Real = PLC AIx_DB.Flow_4.Calibration AT %DB202.DBD734, 1 s

HMI tags "xMotors"
   "Motors_DB_M1_CMD_Hand" : Bool = PLC Motors_DB.M1.CMD.Hand AT %DB204.DBX6.0, 1 s
   "Motors_DB_M1_CMD_Start_M" : Bool = PLC Motors_DB.M1.CMD.Start_M AT %DB204.DBX6.2, 1 s
   "Motors_DB_M1_CMD_Force" : Bool = PLC Motors_DB.M1.CMD.Force AT %DB204.DBX6.3, 1 s
   "Motors_DB_M1_CMD_Service" : Bool = PLC Motors_DB.M1.CMD.Service AT %DB204.DBX6.6, 1 s
   "Motors_DB_M1_CMD_Sim" : Bool = PLC Motors_DB.M1.CMD.Sim AT %DB204.DBX7.2, 1 s
   "Motors_DB_M1_Status" : Int = PLC Motors_DB.M1.Status AT %DB204.DBW10, 1 s
   "Motors_DB_M1_Use_QF" : Bool = PLC Motors_DB.M1.Use.QF AT %DB204.DBX12.1, 1 s
   "Motors_DB_M1_Use_KM" : Bool = PLC Motors_DB.M1.Use.KM AT %DB204.DBX12.2, 1 s
   "Motors_DB_M1_Use_Serivce" : Bool = PLC Motors_DB.M1.Use.Serivce AT %DB204.DBX12.3, 1 s
   "Motors_DB_M1_Use_Termo" : Bool = PLC Motors_DB.M1.Use.Termo AT %DB204.DBX12.4, 1 s
   "Motors_DB_M1_FB_QF" : Bool = PLC Motors_DB.M1.FB.QF AT %DB204.DBX14.1, 1 s
   "Motors_DB_M1_FB_KM" : Bool = PLC Motors_DB.M1.FB.KM AT %DB204.DBX14.2, 1 s
   "Motors_DB_M1_FB_Serivce" : Bool = PLC Motors_DB.M1.FB.Serivce AT %DB204.DBX14.3, 1 s
   "Motors_DB_M1_FB_Termo" : Bool = PLC Motors_DB.M1.FB.Termo AT %DB204.DBX14.4, 1 s
   "Motors_DB_M1_Alarm" : Word = PLC Motors_DB.M1.Alarm AT %DB204.DBW34, 1 s
   "Motors_DB_M1_Res_h" : DInt = PLC Motors_DB.M1.Res_h AT %DB204.DBD36, 1 s
   "Motors_DB_M1_Wait_On_SP" : Int = PLC Motors_DB.M1.Wait_On.SP AT %DB204.DBW18, 1 s
   "Motors_DB_M1_Wait_On_Now" : Int = PLC Motors_DB.M1.Wait_On.Now AT %DB204.DBW20, 1 s
   "Motors_DB_M1_Wait_Off_SP" : Int = PLC Motors_DB.M1.Wait_Off.SP AT %DB204.DBW24, 1 s
   "Motors_DB_M1_Wait_Off_Now" : Int = PLC Motors_DB.M1.Wait_Off.Now AT %DB204.DBW26, 1 s
   "Motors_DB_M2_CMD_Hand" : Bool = PLC Motors_DB.M2.CMD.Hand AT %DB204.DBX50.0, 1 s
   "Motors_DB_M2_CMD_Start_M" : Bool = PLC Motors_DB.M2.CMD.Start_M AT %DB204.DBX50.2, 1 s
   "Motors_DB_M2_CMD_Force" : Bool = PLC Motors_DB.M2.CMD.Force AT %DB204.DBX50.3, 1 s
   "Motors_DB_M2_CMD_Service" : Bool = PLC Motors_DB.M2.CMD.Service AT %DB204.DBX50.6, 1 s
   "Motors_DB_M2_CMD_Sim" : Bool = PLC Motors_DB.M2.CMD.Sim AT %DB204.DBX51.2, 1 s
   "Motors_DB_M2_Status" : Int = PLC Motors_DB.M2.Status AT %DB204.DBW54, 1 s
   "Motors_DB_M2_Use_QF" : Bool = PLC Motors_DB.M2.Use.QF AT %DB204.DBX56.1, 1 s
   "Motors_DB_M2_Use_KM" : Bool = PLC Motors_DB.M2.Use.KM AT %DB204.DBX56.2, 1 s
   "Motors_DB_M2_Use_Serivce" : Bool = PLC Motors_DB.M2.Use.Serivce AT %DB204.DBX56.3, 1 s
   "Motors_DB_M2_Use_Termo" : Bool = PLC Motors_DB.M2.Use.Termo AT %DB204.DBX56.4, 1 s
   "Motors_DB_M2_FB_QF" : Bool = PLC Motors_DB.M2.FB.QF AT %DB204.DBX58.1, 1 s
   "Motors_DB_M2_FB_KM" : Bool = PLC Motors_DB.M2.FB.KM AT %DB204.DBX58.2, 1 s
   "Motors_DB_M2_FB_Serivce" : Bool = PLC Motors_DB.M2.FB.Serivce AT %DB204.DBX58.3, 1 s
   "Motors_DB_M2_FB_Termo" : Bool = PLC Motors_DB.M2.FB.Termo AT %DB204.DBX58.4, 1 s
   "Motors_DB_M2_Alarm" : Word = PLC Motors_DB.M2.Alarm AT %DB204.DBW78, 1 s
   "Motors_DB_M2_Res_h" : DInt = PLC Motors_DB.M2.Res_h AT %DB204.DBD80, 1 s
   "Motors_DB_M2_Wait_On_SP" : Int = PLC Motors_DB.M2.Wait_On.SP AT %DB204.DBW62, 1 s
   "Motors_DB_M2_Wait_On_Now" : Int = PLC Motors_DB.M2.Wait_On.Now AT %DB204.DBW64, 1 s
   "Motors_DB_M2_Wait_Off_SP" : Int = PLC Motors_DB.M2.Wait_Off.SP AT %DB204.DBW68, 1 s
   "Motors_DB_M2_Wait_Off_Now" : Int = PLC Motors_DB.M2.Wait_Off.Now AT %DB204.DBW70, 1 s
   "Motors_DB_M3_CMD_Hand" : Bool = PLC Motors_DB.M3.CMD.Hand AT %DB204.DBX94.0, 1 s
   "Motors_DB_M3_CMD_Start_M" : Bool = PLC Motors_DB.M3.CMD.Start_M AT %DB204.DBX94.2, 1 s
   "Motors_DB_M3_CMD_Force" : Bool = PLC Motors_DB.M3.CMD.Force AT %DB204.DBX94.3, 1 s
   "Motors_DB_M3_CMD_Service" : Bool = PLC Motors_DB.M3.CMD.Service AT %DB204.DBX94.6, 1 s
   "Motors_DB_M3_CMD_Sim" : Bool = PLC Motors_DB.M3.CMD.Sim AT %DB204.DBX95.2, 1 s
   "Motors_DB_M3_Status" : Int = PLC Motors_DB.M3.Status AT %DB204.DBW98, 1 s
   "Motors_DB_M3_Use_QF" : Bool = PLC Motors_DB.M3.Use.QF AT %DB204.DBX100.1, 1 s
   "Motors_DB_M3_Use_KM" : Bool = PLC Motors_DB.M3.Use.KM AT %DB204.DBX100.2, 1 s
   "Motors_DB_M3_Use_Serivce" : Bool = PLC Motors_DB.M3.Use.Serivce AT %DB204.DBX100.3, 1 s
   "Motors_DB_M3_Use_Termo" : Bool = PLC Motors_DB.M3.Use.Termo AT %DB204.DBX100.4, 1 s
   "Motors_DB_M3_FB_QF" : Bool = PLC Motors_DB.M3.FB.QF AT %DB204.DBX102.1, 1 s
   "Motors_DB_M3_FB_KM" : Bool = PLC Motors_DB.M3.FB.KM AT %DB204.DBX102.2, 1 s
   "Motors_DB_M3_FB_Serivce" : Bool = PLC Motors_DB.M3.FB.Serivce AT %DB204.DBX102.3, 1 s
   "Motors_DB_M3_FB_Termo" : Bool = PLC Motors_DB.M3.FB.Termo AT %DB204.DBX102.4, 1 s
   "Motors_DB_M3_Alarm" : Word = PLC Motors_DB.M3.Alarm AT %DB204.DBW122, 1 s
   "Motors_DB_M3_Res_h" : DInt = PLC Motors_DB.M3.Res_h AT %DB204.DBD124, 1 s
   "Motors_DB_M3_Wait_On_SP" : Int = PLC Motors_DB.M3.Wait_On.SP AT %DB204.DBW106, 1 s
   "Motors_DB_M3_Wait_On_Now" : Int = PLC Motors_DB.M3.Wait_On.Now AT %DB204.DBW108, 1 s
   "Motors_DB_M3_Wait_Off_SP" : Int = PLC Motors_DB.M3.Wait_Off.SP AT %DB204.DBW112, 1 s
   "Motors_DB_M3_Wait_Off_Now" : Int = PLC Motors_DB.M3.Wait_Off.Now AT %DB204.DBW114, 1 s
